// Mitsubishi GX Works2 project: ZhaoQing_HuaCheng1_Debug   PLC: Q06UDEH (continued)

H1000Conveyor7(ConveyorMotor:=H1000Conveyor7IO);
H1000Conveyor7IO.xForward:=M66;
H1000Conveyor7IO.xCWPresent:=X4F;
Y14F:=H1000Conveyor7IO.xMotorCW;
H1000Conveyor7IO.iDeviceID:=1007;

H1000Conveyor8(ConveyorMotor:=H1000Conveyor8IO);
H1000Conveyor8IO.xForward:=M67;
H1000Conveyor8IO.xCWPresent:=X50;
Y150:=H1000Conveyor8IO.xMotorCW;
H1000Conveyor8IO.iDeviceID:=1008;

H1000Conveyor9(ConveyorMotor:=H1000Conveyor9IO);
H1000Conveyor9IO.xForward:=M68;
H1000Conveyor9IO.xCWPresent:=X51;
Y151:=H1000Conveyor9IO.xMotorCW;
H1000Conveyor9IO.iDeviceID:=1009;

H1000Conveyor10(ConveyorMotor:=H1000Conveyor10IO);
H1000Conveyor10IO.xForward:=M67;
H1000Conveyor10IO.xCWPresent:=X52;
Y152:=H1000Conveyor10IO.xMotorCW;
H1000Conveyor10IO.iDeviceID:=1010;
(*注液隔离仓*)
(*FillQuarantineDoorInside(ShuttleCarInOut:= FillQuarantineDoorInsideIO );
FillQuarantineDoorInsideIO.xCylinder:=1;
ShuttleCarCurrentPosition(X109 OR X10A ,X10A ,X109, FALSE,FillQuarantineDoorInsideIO.iCurrentPos);
FillQuarantineDoorInsideIO.xForward:=M191;
FillQuarantineDoorInsideIO.xBackward:=M192 ;
Y160:=FillQuarantineDoorInsideIO.xCW;
Y161:=FillQuarantineDoorInsideIO.xCCW;

FillQuarantineDoorOutside(ShuttleCarInOut:= FillQuarantineDoorOutsideIO );
FillQuarantineDoorOutsideIO.xCylinder:=1;
ShuttleCarCurrentPosition(X10B OR X10C ,X10C ,X10B, FALSE,FillQuarantineDoorOutsideIO.iCurrentPos);
FillQuarantineDoorOutsideIO.xForward:=M193;
FillQuarantineDoorOutsideIO.xBackward:=M194 ;
Y162:=FillQuarantineDoorOutsideIO.xCW;
Y163:=FillQuarantineDoorOutsideIO.xCCW;*)
(*注液入与出线体*)
H850Conveyor1(ConveyorMotor:=H850Conveyor1IO);
H850Conveyor1IO.xForward:=M129;
H850Conveyor1IO.xCWPresent:=X78;
Y178:=H850Conveyor1IO.xMotorCW;
H850Conveyor1IO.iDeviceID:=8501;

H850Conveyor3(ConveyorMotor:=H850Conveyor3IO);
H850Conveyor3IO.xForward:=M130;
H850Conveyor3IO.xCWPresent:=X7A;
Y17A:=H850Conveyor3IO.xMotorCW;
H850Conveyor3IO.iDeviceID:=8503;

H850Conveyor4(ConveyorMotor:=H850Conveyor4IO);
H850Conveyor4IO.xForward:=M131;
H850Conveyor4IO.xCWPresent:=X7B;
Y17B:=H850Conveyor4IO.xMotorCW;
H850Conveyor4IO.iDeviceID:=8504;

H850Conveyor5(ConveyorMotor:=H850Conveyor5IO);
H850Conveyor5IO.xForward:=M132;
H850Conveyor5IO.xCWPresent:=X7C;
Y17C:=H850Conveyor5IO.xMotorCW;
H850Conveyor5IO.iDeviceID:=8505;

H850Conveyor6(ConveyorMotor:=H850Conveyor6IO);
H850Conveyor6IO.xForward:=M133;
H850Conveyor6IO.xCWPresent:=X7D;
Y17D:=H850Conveyor6IO.xMotorCW;
H850Conveyor6IO.iDeviceID:=8506;

H850Conveyor7(ConveyorMotor:=H850Conveyor7IO);
H850Conveyor7IO.xForward:=M164;
H850Conveyor7IO.xCWPresent:=X7E;
Y17E:=H850Conveyor7IO.xMotorCW;
H850Conveyor7IO.iDeviceID:=8507;

H850Rotor(ShuttleCarInOut:=H850RotorIO);
ShuttleCarCurrentPosition(X82 OR X76  ,X82 ,X76, FALSE,H850RotorIO.iCurrentPos);
H850RotorIO.xReady:=TRUE;
H850RotorIO.xForward:=M75;
H850RotorIO.xBackward:=M76;
H850RotorIO.xPosLimit:=X84;
H850RotorIO.xNegLimit:=X85;
Y182:=H850RotorIO.xCW;
Y183:=H850RotorIO.xCCW;
Y1B9:=H850RotorIO.xBrake;

H850RotorConveyor(ConveyorMotor:=H850RotorConveyorIO);
H850RotorConveyorIO.xForward:=M77;
H850RotorConveyorIO.xBackward:=M82;
H850RotorConveyorIO.xCWPresent:=X87;
H850RotorConveyorIO.xCCWPresent:=X86;
Y185:=H850RotorConveyorIO.xMotorCW;
Y184:=H850RotorConveyorIO.xMotorCCW;
H850RotorConveyorIO.xUnloadCCW:=1;
H850RotorConveyorIO.tLoadDelay:=T#2s;
H850RotorConveyorIO.iDeviceID:=8599;

H850Switch(ConveyorEntryIO:=H850SwitchConveyorIn,ConveyorExitIO:=H850SwitchConveyorOut,SwitchIO:=H850SwitchIO);
H850SwitchIO.xLiftCylinderExtendButton:=M71;
H850SwitchIO.xLiftCylinderRetractButton:=M72;
Y189:=H850SwitchIO.xLiftCylinderExtend;
Y188:=H850SwitchIO.xLiftCylinderRetract;
H850SwitchIO.xLiftCylinderExtendDetect:=X88;
H850SwitchIO.xLiftCylinderRetractDetect:=X89;
H850SwitchConveyorIn.xForward:=M70;
H850SwitchConveyorIn.xCWPresent:=XB4;
Y19B:=H850SwitchConveyorIn.xMotorCW;
Y139:=H850SwitchConveyorIn.xMotorCW;(*新加的滚轮电机*)
H850SwitchConveyorIn.tLoadDelay:=T#2s;
H850SwitchConveyorIn.iDeviceID:=8598;
H850SwitchConveyorOut.xForward:=M73;
H850SwitchConveyorOut.xCWPresent:=X8A;
Y18A:=H850SwitchConveyorOut.xMotorCW;
H850SwitchConveyorOut.iDeviceID:=8598;


H850Conveyor8(ConveyorMotor:=H850Conveyor8IO);
H850Conveyor8IO.xForward:=M74;
H850Conveyor8IO.xCWPresent:=X7F;
Y17F:=H850Conveyor8IO.xMotorCW;
H850Conveyor8IO.iDeviceID:=8508;
(*高温库前线体*)
(*-------高温入库分流扫码*)
IF X0BB AND NOT X0BA  THEN 
	Y1BE:=0;
	Y1BF:=1;
END_IF ;
IF ldp(TRUE,X0BA AND D2300=0)  THEN 
	Y1BE:=0;
	Y1BF:=0;
	xscaning1:=1;
END_IF ;
IF ldp(TRUE, D2300=2 OR D2300=3) THEN
	Y1BE:=1;
    Y1BF:=1;
    xscaning1:=0;
END_IF;  
(*阻挡气缸升起，检测有无信号存在，上位机扫码信号复位，可以扫码*)
IF X0BA AND D2300=0 AND Y1BE = 0 AND Y1BF=0 THEN 
	D3300:=2;
END_IF;
(*单体复位后把扫码信息复位*)
IF g_xResetSingle AND g_iDeviceIDSelect=H2200Switch2ConveyorIn.iDeviceID THEN
	xscaning1:=0;
	D3300:=1;
END_IF;
IF D2300 =1 AND g_xReset THEN(*扫码失败复位*)
	D3300:=0;
END_IF;
(* 顶升移载收到物料后复位读码信号*)
(*IF LDP(TRUE,Import1SwitchConveyorOut.xEmpty=0 AND D2300=2) OR LDP(TRUE,Import2SwitchConveyorOut.xEmpty=0 AND D2300=3) THEN*)
	(*修改下复位扫码的时序，分流后再复位扫码信息，方便分流*)
IF( Import1Conveyor1IO.xEmpty=0 AND D2300=2) OR  (Import2Conveyor1IO.xEmpty=0 AND D2300=3) THEN(*效率低*)(*效率低也没办法，分流信息不能提前复位*)
(*IF (Import1SwitchConveyorOut.xBusy AND D2300=2) OR (Import2SwitchConveyorOut.xBusy AND D2300=3) THEN*)
	D3300:=1;    (*接堆垛机那个口顶起来才允许下一次扫码*)(*到达分流顶升移载后复位*)
END_IF;
	(*------高温出库分流扫码*)
	IF X106 THEN 
	xScaning2:=0;
END_IF;
IF X0B9 AND NOT X0B8  THEN 
	Y1BC:=0;
	Y1BD:=1;
END_IF ;
IF X0B8 AND  D2305=0  THEN 
	Y1BC:=0;
	Y1BD:=0;
	xScaning2:=1;
END_IF ;
IF ldp(TRUE,  D2305=2 OR D2305=3) THEN
	Y1BC:=1;
    Y1BD:=1;
    xScaning2:=0;
END_IF;
IF X0B8  AND D2305=0 THEN 
	D3305:=2;
END_IF;
IF X2F OR X39 OR g_xReset THEN(*增加复位信号，扫码失败后按复位按钮*)
	D3305:=1;(*运出之后才允许下一次扫码*)
	END_IF;
(*1巷道入库*)
Import1Conveyor1(ConveyorMotor:=Import1Conveyor1IO);
Import1Conveyor1IO.xForward:=M98;
Import1Conveyor1IO.xCWPresent:=XE3;
Y1F4:=Import1Conveyor1IO.xMotorCW;
Import1Conveyor1IO.iDeviceID:=2290;

Import1Conveyor2(ConveyorMotor:=Import1Conveyor2IO);
Import1Conveyor2IO.tLoadDelay:=T#1s;
Import1Conveyor2IO.xForward:=M99;
Import1Conveyor2IO.xCWPresent:=XE4;
Y1F5:=Import1Conveyor2IO.xMotorCW;
Import1Conveyor2IO.iDeviceID:=2289;

Import1Switch(ConveyorEntryIO:=Import1SwitchConveyorIn,
                          ConveyorExitIO:=Import1SwitchConveyorOut ,
                           SwitchIO:=Import1SwitchIO);
Import1SwitchIO.xLiftCylinderExtendButton:=M147;
Import1SwitchIO.xLiftCylinderRetractButton:=M148;
Import1SwitchIO.xExitBarCylinderRetractButton:=M161;
Y1E0:=Import1SwitchIO.xExitBarCylinderRetract;
Y1E2:=Import1SwitchIO.xLiftCylinderExtend;
Y1E1:=Import1SwitchIO.xLiftCylinderRetract;
Import1SwitchIO.xLiftCylinderExtendDetect:=XE1;
Import1SwitchIO.xLiftCylinderRetractDetect:=XE2; 
Import1SwitchConveyorIn.xCWPresent:=XE0;
Import1SwitchConveyorIn.tLoadDelay:=T#3s;
Import1SwitchConveyorIn.iDeviceID:=2297;
Import1SwitchConveyorOut.xForward:=M149;
Import1SwitchConveyorOut.xCWPresent:=X108;
Y1F6:=Import1SwitchConveyorOut.xMotorCW;
Import1SwitchConveyorOut.iDeviceID:=2297;

Import1LoadCylinder(ShuttleCarInOut:=Import1LoadCylinderIO);
ShuttleCarCurrentPosition(XE7 OR XE6,XE7 ,XE6, FALSE,Import1LoadCylinderIO.iCurrentPos );
Import1LoadCylinderIO.xReady:=TRUE;
Import1LoadCylinderIO.xForward:=M159;
Import1LoadCylinderIO.xBackward:=M160;
Import1LoadCylinderIO.xPosLimit:=TRUE;
Import1LoadCylinderIO.xNegLimit:=TRUE;
Y1E4:=Import1LoadCylinderIO.xCW;
Y1E3:=Import1LoadCylinderIO.xCCW;

(*1巷道出库*)
Export1Conveyor1(ConveyorMotor:=Export1Conveyor1IO);
Export1Conveyor1IO.xForward:=M94;
Export1Conveyor1IO.xCWPresent:=XEC;
Y1F7:=Export1Conveyor1IO.xMotorCW;
Export1Conveyor1IO.iDeviceID:=3081;

Export1Conveyor2(ConveyorMotor:=Export1Conveyor2iO);
Export1Conveyor2IO.xForward:=M95;
Export1Conveyor2IO.xCWPresent:=XEB;
Y1F8:=Export1Conveyor2IO.xMotorCW;
Export1Conveyor2IO.iDeviceID:=3082;

Export1Switch(ConveyorEntryIO:=Export1SwitchConveyorIn,
                          ConveyorExitIO:=Export1SwitchConveyorOut ,
                           SwitchIO:=Export1SwitchIO);
Export1SwitchIO.xLiftCylinderExtendButton:=M150;
Export1SwitchIO.xLiftCylinderRetractButton:=M151;
Y1E7:=Export1SwitchIO.xLiftCylinderExtend;
Y1E6:=Export1SwitchIO.xLiftCylinderRetract;
Export1SwitchIO.xLiftCylinderExtendDetect:=XE9;
Export1SwitchIO.xLiftCylinderRetractDetect:=XEA;
Export1SwitchConveyorIn.xForward:=M152;
Export1SwitchConveyorIn.xCWPresent:=X106;
Export1SwitchConveyorIn.tLoadDelay:=T#2s;
Export1SwitchConveyorIn.iDeviceID:=3083;
Y1F9:=Export1SwitchConveyorIn.xMotorCW;
Export1SwitchConveyorOut.xCWPresent:=X106;
Export1SwitchConveyorOut.iDeviceID:=3083;

Export1LoadCylinder(ShuttleCarInOut:=Export1LoadCylinderIO);
ShuttleCarCurrentPosition(XEF OR XEE ,XEF ,XEE, FALSE,Export1LoadCylinderIO.iCurrentPos);
Export1LoadCylinderIO.xReady:=TRUE;
Export1LoadCylinderIO.xForward:=M157;
Export1LoadCylinderIO.xBackward:=M158;
Export1LoadCylinderIO.xPosLimit:=TRUE;
Export1LoadCylinderIO.xNegLimit:=TRUE;
Y1E9:=Export1LoadCylinderIO.xCW;
Y1E8:=Export1LoadCylinderIO.xCCW;


(*2巷道入库*)
Import2Conveyor1(ConveyorMotor:=Import2Conveyor1IO);
Import2Conveyor1IO.xForward:=M153;
Import2Conveyor1IO.xCWPresent:=XF3;
Y1FA:=Import2Conveyor1IO.xMotorCW;
Import2Conveyor1IO.iDeviceID:=2288;

Import2Conveyor2(ConveyorMotor:=Import2Conveyor2IO);
Import2Conveyor2IO.tLoadDelay:=T#1s;
Import2Conveyor2IO.xForward:=M154;
Import2Conveyor2IO.xCWPresent:=XF4;
Y1FB:=Import2Conveyor2IO.xMotorCW;
Import2Conveyor2IO.iDeviceID:=2287;

Import2Switch(ConveyorEntryIO:=Import2SwitchConveyorIn,
                          ConveyorExitIO:=Import2SwitchConveyorOut ,
                           SwitchIO:=Import2SwitchIO);
Import2SwitchIO.xLiftCylinderExtendButton:=M155;
Import2SwitchIO.xLiftCylinderRetractButton:=M156;
Y1EC:=Import2SwitchIO.xLiftCylinderExtend;
Y1EB:=Import2SwitchIO.xLiftCylinderRetract;
Import2SwitchIO.xLiftCylinderExtendDetect:=XF1;
Import2SwitchIO.xLiftCylinderRetractDetect:=XF2;
Import2SwitchConveyorIn.xCWPresent:=X104;
Import2SwitchConveyorIn.tLoadDelay:=T#2s;
Import2SwitchConveyorIn.iDeviceID:=2296;
Import2SwitchConveyorOut.xForward:=M165;
Import2SwitchConveyorOut.xCWPresent:=X100;
Y1FC:=Import2SwitchConveyorOut.xMotorCW;
Import2SwitchConveyorOut.iDeviceID:=2296;

Import2LoadCylinder(ShuttleCarInOut:=Import2LoadCylinderIO);
ShuttleCarCurrentPosition(XF6 OR XF7 ,XF7 ,XF6, FALSE,Import2LoadCylinderIO.iCurrentPos );
Import2LoadCylinderIO.xReady:=TRUE;
Import2LoadCylinderIO.xForward:=M171;
Import2LoadCylinderIO.xBackward:=M162;
Import2LoadCylinderIO.xPosLimit:=TRUE;
Import2LoadCylinderIO.xNegLimit:=TRUE;
Y1EE:=Import2LoadCylinderIO.xCW;
Y1ED:=Import2LoadCylinderIO.xCCW;

(*2巷道出库*)
Export2Conveyor1(ConveyorMotor:=Export2Conveyor1IO);
Export2Conveyor1IO.xForward:=M96;
Export2Conveyor1IO.xCWPresent:=XFB;
Y1FD:=Export2Conveyor1IO.xMotorCW;
Export2Conveyor1IO.iDeviceID:=3085;

Export2Conveyor2(ConveyorMotor:=Export2Conveyor2iO);
Export2Conveyor2IO.xForward:=M97;
Export2Conveyor2IO.xCWPresent:=XFC;
Y1FE:=Export2Conveyor2IO.xMotorCW;
Export2Conveyor2IO.iDeviceID:=3086;

Export2Switch(ConveyorEntryIO:=Export2SwitchConveyorIn,
                          ConveyorExitIO:=Export2SwitchConveyorOut ,
                           SwitchIO:=Export2SwitchIO);
Export2SwitchIO.xLiftCylinderExtendButton:=M120;
Export2SwitchIO.xLiftCylinderRetractButton:=M121;
Export2SwitchIO.xLiftCylinderExtendInit:=1;
Y1F1:=Export2SwitchIO.xLiftCylinderExtend;
Y1F0:=Export2SwitchIO.xLiftCylinderRetract;
Export2SwitchIO.xLiftCylinderExtendDetect:=XF9;
Export2SwitchIO.xLiftCylinderRetractDetect:=XFA;
Export2SwitchConveyorIn.xForward:=M123;
Export2SwitchConveyorIn.xCWPresent:=X105;
Export2SwitchConveyorIn.tLoadDelay:=T#2s;
Y1FF:=Export2SwitchConveyorIn.xMotorCW;
Export2SwitchConveyorIn.iDeviceID:=3084;
Export2SwitchConveyorOut.xCWPresent:=X105;
Export2SwitchConveyorOut.iDeviceID:=3084;

Export2LoadCylinder(ShuttleCarInOut:=Export2LoadCylinderIO);
ShuttleCarCurrentPosition( XFF OR XFE ,XFF ,XFE, FALSE, Export2LoadCylinderIO.iCurrentPos);
Export2LoadCylinderIO.xReady:=TRUE;
Export2LoadCylinderIO.xForward:=M124;
Export2LoadCylinderIO.xBackward:=M125;
Export2LoadCylinderIO.xPosLimit:=TRUE;
Export2LoadCylinderIO.xNegLimit:=TRUE;
Y1F2:=Export2LoadCylinderIO.xCW;
Y1F3:=Export2LoadCylinderIO.xCCW;




IF g_xAuto THEN
	(**高温库前自动程序**)
	Y1EA:=1;
	m_tonScan2(IN:=xScaning2 ,PT:=T#500ms ,Q:=m_xScan2,ET:= m_tScan2 );(*---------扫码标志位做延时，防止走不到位*)
	Y187:=NOT m_xScan2 AND  m_iExportConveyorOcuppy<>0;(***出库倍速链***)(*---------扫码时停下，扫完走*)
	Y1BA:=NOT m_xScan2 AND  m_iExportConveyorOcuppy<>0;(*后增加滚筒线，在出库线占用状态字有的情况下开始旋转*)
	Y19E :=NOT m_xScan2 AND  m_iExportConveyorOcuppy<>0;
	Y19F:=NOT m_xScan2 AND  m_iExportConveyorOcuppy<>0; 
	(**高温库1巷道出库**)
	(*************************
	上位机通讯程序3
	出口状态  D3105
	1:禁止出库
    2:允许出库
    
    1线堆积(化成线)状态	3106	"1：正常2:堆积 "

2线(二封线)堆积状态	3107	"1：正常2:堆积 "


    收到空框请求D2105
    1：复位，
    2：收到出库请求
	**********************出库********************************)
	(******1巷道******)
	IF NOT XED  AND NOT XEB AND NOT Y1F8 AND Export1LoadCylinderIO.iCurrentPos=2 THEN(*-----这里加了很多条件，保证不会轻易顶起来*)
		D3105:=2;
	ELSE
		D3105:=1;
	END_IF;
	m_tonHangUpChemDalay(IN:= H2200Conveyor5IO.xEmpty=0 OR H2200Conveyor6IO.xEmpty=0  ,PT:=T#30S ,Q:= m_xHangUpChem,ET:= m_tHangUpChemDalayCurrentTime );
	m_tonHangUpPackageDalay(IN:= H3000Conveyor9IO.xEmpty=0 OR H3000Conveyor10IO.xEmpty=0 ,PT:=T#10S ,Q:= m_xHangUpPackage,ET:= m_tHangUpPackageDalayCurrentTime );
	IF m_xHangUpChem THEN
		D3106:=2;
		D3126:=2;
	ELSE
		D3106:=1;
		D3126:=1;
	END_IF;
	
	IF m_xHangUpPackage THEN
		D3107:=2;
		D3127:=2;
	ELSE
		D3107:=1;
		D3127:=1;
	END_IF;
	
	IF D2105=2 THEN
		M883:=1;
	ELSE
		M883:=0;
	END_IF;
	(******2巷道******)
   (*************************
	上位机通讯程序
	出口状态  D3125
	1:禁止出库
    2:允许出库
    1线堆积(化成线)状态	3126	"1：正常2:堆积 "
2线(二封线)堆积状态	3127	"1：正常2:堆积 "

    收到空框请求D2125
    1：复位，
    2：收到出库请求
	**********************出库********************************)
	IF NOT XFD AND Export2LoadCylinderIO.iCurrentPos=2 THEN
		D3125:=2;
	ELSE
		D3125:=1;
	END_IF;
	IF D2125=2 THEN
		M884:=1;
	ELSE
		M884:=0;
	END_IF;
	(*********************入库****************************)
	(***********************************
	入口状态 D3100
	1:无电池入库请求
     2:有电池入库请求
	************************************)
	(******1巷道******)
	m_tonImport1RequestDalay(IN:= XE5 ,PT:= t#3S ,Q:= m_xImport1RequestDalay ,ET:=m_tImport1RequestDalaDalayCurren);
	IF m_xImport1RequestDalay AND Import1LoadCylinderIO.iCurrentPos=2 THEN
		D3100:=2;
	ELSE
		D3100:=1;
    END_IF;  
    (******2巷道******)
	m_tonImport2RequestDalay(IN:= XF5 ,PT:= t#3S ,Q:= m_xImport2RequestDalay ,ET:=m_tImport2RequestDalaDalayCurren);    
    IF m_xImport2RequestDalay  AND Import2LoadCylinderIO.iCurrentPos=2 THEN
		D3120:=2;
	ELSE
		D3120:=1;
    END_IF;
    (*******************************************************)
    (******高温出库分流******)
    (***********************************
	有板状态 D3305
	1：无板，2：有板
    分流方向 D2305
0：复位
1：读码失败
2：满筐进加压化成
3：满筐进二封
4：空筐回流进注液
	************************************)
	(*IF H3000SwitchPackageConveyorIn.xEmpty=0 THEN
		D3305:=1;
	ELSE
		D3305:=2;
	END_IF;*)
	IF D2305=2 THEN
		M882:=1;
	END_IF;
	IF D2305 =3 THEN
		M882:=0;
	END_IF;
	(**********************************)
	 (******高温出库后升降机2分流******)
	     (***********************************
	有板状态 D3310
	1：无板，2：有板
    分流方向 D2310
0：复位
1：读码失败
2：空筐去注液
3：满筐去加压化成
	************************************)
	IF X3B THEN
		D3310:=2;
	ELSE
		D3310:=1;
	END_IF;
	(*
	IF D2310=2 THEN        ------------这段屏蔽了，直接加到xcondition里了
        Lifter2ExportChem:=01;
	END_IF;
	IF D2310=3 THEN
        Lifter2ExportChem:=1;
	END_IF;
	*)
	(*************	"化成后站台40082335	5	
	分流方向	2335	"0：复位
1：读码失败
2：处理完成放行"
"**********************)



	IF H1000Conveyor2IO.xEmpty=0 THEN
		D3335:=2;
	ELSE
		D3335:=1;
	END_IF;
	IF NOT H850Conveyor8IO.xEmpty THEN
		D3340:=2;
	ELSE
		D3340:=1;
		END_IF;
  (***********************************)
	IF  LDP(TRUE,M883) AND XED THEN
        Export1LoadCylinderIO.xMDIExe:=1;
        Export1LoadCylinderIO.iDestinationPos:=1;
	END_IF;
	IF NOT XED AND NOT XEB  AND NOT Y1F8 AND  Export1Conveyor2IO.xEmpty AND NOT Export1Conveyor2IO.xBusy THEN
        Export1LoadCylinderIO.xMDIExe:=1;
        Export1LoadCylinderIO.iDestinationPos:=2;
     END_IF;		
	Export1Conveyor2IO.xLoad:=XED AND Export1LoadCylinderIO.iCurrentPos=1;
	Export1Conveyor2IO.xUnload:=Export1Conveyor1IO.xEmpty;
	Export1Conveyor1IO.xLoad:=Export1Conveyor2IO.xNextRun;

	Export1Conveyor1Io.xUnload:=Export1SwitchConveyorIn.xEmpty  AND  m_iExportConveyorOcuppy=1 AND  NOT M173;
	IF Export1Conveyor1Io.xEmpty=0 AND m_xExportConveyorIdle THEN
		m_iExportConveyorOcuppy:=1;
	END_IF;
	Export1SwitchIO.xEntryEnable:=Export1Conveyor1Io.xNextRun;
	Export1SwitchIO.xSwithEnable:=1;
	(*倍速链上只有一个物料出库*)
   Export1SwitchIO.xExitEnable:=(H3000SwitchChemConveyorIn.xEmpty AND M882) OR (H3000Conveyor1IO.xEmpty AND NOT M882);
	(**高温库2巷道出库**)
	IF  LDP(TRUE,M884) AND XFD THEN
        Export2LoadCylinderIO.xMDIExe:=1;
        Export2LoadCylinderIO.iDestinationPos:=1;
	END_IF;
	IF NOT XFD  AND NOT Export2Conveyor1IO.xBusy AND Export2Conveyor1IO.xEmpty  THEN
        Export2LoadCylinderIO.xMDIExe:=1;
        Export2LoadCylinderIO.iDestinationPos:=2;
     END_IF;	
	Export2Conveyor1IO.xLoad:=XFD AND Export2LoadCylinderIO.iCurrentPos=1;
	Export2Conveyor1IO.xUnload:=Export2Conveyor2IO.xEmpty;
	Export2Conveyor2IO.xLoad:=Export2Conveyor1IO.xNextRun;
(*	Export2Conveyor2Io.xUnload:=Export2SwitchConveyorIn.xEmpty AND NOT XE8 AND NOT Y1E5;(*增加阻挡器信号与到位信号*)
	Export2Conveyor2Io.xUnload:=Export2SwitchConveyorIn.xEmpty AND  m_iExportConveyorOcuppy=2 AND NOT M173;
	Export2SwitchIO.xEntryEnable:=Export2Conveyor2Io.xNextRun;
	Export2SwitchIO.xSwithEnable:=1;

	IF Export2Conveyor2Io.xEmpty=0 AND m_xExportConveyorIdle  THEN
		m_iExportConveyorOcuppy:=2;
	END_IF;
	IF m_iExportConveyorOcuppy=2  THEN
		Y1E5:=1;(*1巷道出库阻挡器*)
		Export1SwitchIO.xLiftCylinderExtendInit:=0;
	ELSE
		Y1E5:=0;(*1巷道出库阻挡器*)
		Export1SwitchIO.xLiftCylinderExtendInit:=1;	
	END_IF;
	
	Export2SwitchIO.xExitEnable:=(H3000SwitchChemConveyorIn.xEmpty AND M882) OR (H3000Conveyor1IO.xEmpty AND NOT M882);
	(*占用信号的复位*)
	IF LDP(TRUE,H3000SwitchChemConveyorIn.xEmpty=0 AND M882) OR LDP(TRUE,H3000Conveyor1IO.xEmpty=0 AND NOT M882) THEN
		m_iExportConveyorOcuppy:=0;
	END_IF;
	
	m_tonExportConveyorOcuppy(IN:= m_iExportConveyorOcuppy=0 ,PT:= T#3s ,Q:= m_xExportConveyorIdle ,ET:= m_tExportConveyorOcuppyCurrent );

	(*满框出库去二次封装线体*)
	H3000SwitchQuadPackageIO.xEntryEnable:=1;(*这里要加扫码条件*)
	H3000SwitchQuadPackageIO.xSwithEnable:= NOT M882;(*触摸屏上按钮选择去化成还是去二封，后期通过上位机扫码给出*)
	IF H3000SwitchQuadPackageIO.xSwithEnable THEN
		H3000SwitchQuadPackageio.xExitEnable:=H3000Conveyor1IO.xEmpty;
		H3000Conveyor1Io.xLoad:=H3000SwitchPackageConveyorOut.xNextRun;
	ELSE
		H3000SwitchQuadPackageio.xExitEnable:=0;	
		H3000Conveyor1Io.xLoad:=0;
	END_IF;
	H3000Conveyor1IO.xUnload:=H3000Conveyor2IO.xEmpty;
	H3000Conveyor2IO.xLoad:=H3000Conveyor1IO.xNextRun;
	H3000Conveyor2IO.xUnload:=H3000Conveyor3IO.xEmpty;
	H3000Conveyor3IO.xLoad:=H3000Conveyor2IO.xNextRun;	
	H3000Conveyor3IO.xUnload:=H3000Conveyor4IO.xEmpty;
	H3000Conveyor4IO.xLoad:=H3000Conveyor3IO.xNextRun;
	H3000Conveyor4IO.xUnload:=H3000Conveyor5IO.xEmpty;
	H3000Conveyor5IO.xLoad:=H3000Conveyor4IO.xNextRun;
	H3000Conveyor5IO.xUnload:=H3000Conveyor6IO.xEmpty;
	H3000Conveyor6IO.xLoad:=H3000Conveyor5IO.xNextRun;
	H3000Conveyor6IO.xUnload:=H3000Conveyor7IO.xEmpty;
	H3000Conveyor7IO.xLoad:=H3000Conveyor6IO.xNextRun;
	H3000Conveyor7IO.xUnload:=H3000Conveyor8IO.xEmpty;
	H3000Conveyor8IO.xLoad:=H3000Conveyor7IO.xNextRun;	
	H3000Conveyor8IO.xUnload:=H3000Conveyor9IO.xEmpty;
	H3000Conveyor9IO.xLoad:=H3000Conveyor8IO.xNextRun;	
	H3000Conveyor9IO.xUnload:=H3000Conveyor10IO.xEmpty;
	H3000Conveyor10IO.xLoad:=H3000Conveyor9IO.xNextRun;
	H3000Conveyor10IO.xUnload:=D401.0;
	D201.0:=H3000Conveyor10IO.xNextRun;
    (**满框去化成**)
	H3000SwitchChemIO.xEntryEnable:=1;
	H3000SwitchChemIO.xSwithEnable:=1;
	H3000SwitchChemIO.xExitEnable:=H3000ChemConveyor2IO.xEmpty;
	H3000SwitchPackageConveyorIn.xUnload:=H3000SwitchChemConveyorIn.xEmpty;
	H3000ChemConveyor2IO.xLoad:=H3000SwitchChemConveyorOut.xNextRun;
	H3000ChemConveyor2IO.xUnload:=H3000ChemConveyor3IO.xEmpty;
	H3000ChemConveyor3IO.xLoad:=H3000ChemConveyor2IO.xNextRun;
	(*临时程序，Lifter2ExportChem:=1;以后要考虑空框回注液的程序，上位机扫码后判断是满框去化成还是空框去注液*)
	IF H3000ChemConveyor3IO.xEmpty=0 AND ( Lifter2TaskID=3 OR Lifter2TaskID=4)  THEN(*这里加扫码成功条件*)
		Lifter2IO.xMDIExe:=1;
		Lifter2IO.iDestinationPos:=5;
	END_IF;
	IF Lifter2IO.iCurrentPos=5 AND abs(D190-Lifter2Position[Lifter2IO.iDestinationPos])<20 AND (Lifter2TaskID=3 OR Lifter2TaskID=4)   THEN	
        Conveyor2IO.xLoad:=H3000ChemConveyor3IO.xNextRun;
        H3000ChemConveyor3IO.xUnload:=Conveyor2IO.xEmpty AND H2200Conveyor1io.xEmpty;(*-------这里防止东西堵在车上*)
         Conveyor2IO.xloadCCW:=0;
	ELSE
		H3000ChemConveyor3IO.xUnload:=0;
	END_IF; 
	   IF Conveyor2IO.xEmpty=0 AND Lifter2TaskID=3 THEN
	   		Lifter2IO.xMDIExe:=1;
			Lifter2IO.iDestinationPos:=4;
	   END_IF;
	   	   IF Conveyor2IO.xEmpty=0 AND Lifter2TaskID=4 THEN
	   		Lifter2IO.xMDIExe:=1;
			Lifter2IO.iDestinationPos:=3;
	   END_IF;
	 IF Lifter2IO.iCurrentPos=4 AND abs(D190-Lifter2Position[Lifter2IO.iDestinationPos])<=20  THEN	
	 	H2200Conveyor1IO.xLoad:=Conveyor2IO.xNextRun; 
	 	Conveyor2IO.xUnload:=H2200Conveyor1IO.xEmpty;
	 	Conveyor2IO.xUnloadCCW:=0;
	 ELSE
	 	H2200Conveyor1IO.xLoad:=0;
	 END_IF;  
	      
	H2200Conveyor1IO.xUnload:=H2200Conveyor2IO.xEmpty;
	H2200Conveyor2IO.xLoad:=H2200Conveyor1IO.xNextRun;
	H2200Conveyor2IO.xUnload:=H2200Conveyor3IO.xEmpty;
	H2200Conveyor3IO.xLoad:=H2200Conveyor2IO.xNextRun;	
	H2200Conveyor3IO.xUnload:=H2200Conveyor4IO.xEmpty;
	H2200Conveyor4IO.xLoad:=H2200Conveyor3IO.xNextRun;
	H2200Conveyor4IO.xUnload:=H2200Conveyor5IO.xEmpty;
	H2200Conveyor5IO.xLoad:=H2200Conveyor4IO.xNextRun;
	H2200Conveyor5IO.xUnload:=H2200Conveyor6IO.xEmpty;
	H2200Conveyor6IO.xLoad:=H2200Conveyor5IO.xNextRun;
	H2200Conveyor6IO.xUnload:=H2200Conveyor7IO.xEmpty;
	H2200Conveyor7IO.xLoad:=H2200Conveyor6IO.xNextRun;
	H2200Conveyor7IO.xUnload:=H2200Conveyor8IO.xEmpty;
	H2200Conveyor8IO.xLoad:=H2200Conveyor7IO.xNextRun;	
	H2200Conveyor8IO.xUnload:=H2200Conveyor9IO.xEmpty;
	H2200Conveyor9IO.xLoad:=H2200Conveyor8IO.xNextRun;	
	H2200Conveyor9IO.xUnload:=H2200Conveyor10IO.xEmpty;
	H2200Conveyor10IO.xLoad:=H2200Conveyor9IO.xNextRun;
	H2200Conveyor10IO.xUnload:=D401.1;
	D201.1:=H2200Conveyor10IO.xNextRun;
	(*化成回流线体*)
	D201.2:=H1000Conveyor10IO.xEmpty;
	H1000Conveyor10IO.xLoad:=D401.2;
	H1000Conveyor10IO.xUnload:=H1000Conveyor9IO.xEmpty;
    H1000Conveyor9IO.xLoad:=H1000Conveyor10IO.xNextRun;
    H1000Conveyor9IO.xUnload:=H1000Conveyor8IO.xEmpty;
    H1000Conveyor8IO.xLoad:=H1000Conveyor9IO.xNextRun;
    H1000Conveyor8IO.xUnload:=H1000Conveyor7IO.xEmpty;
    H1000Conveyor7IO.xLoad:=H1000Conveyor8IO.xNextRun;
    H1000Conveyor7IO.xUnload:=H1000Conveyor6IO.xEmpty;
    H1000Conveyor6IO.xLoad:=H1000Conveyor7IO.xNextRun;
    H1000Conveyor6IO.xUnload:=H1000Conveyor5IO.xEmpty;
    H1000Conveyor5IO.xLoad:=H1000Conveyor6IO.xNextRun;
    H1000Conveyor5IO.xUnload:=H1000Conveyor4IO.xEmpty;
    H1000Conveyor4IO.xLoad:=H1000Conveyor5IO.xNextRun;
    H1000Conveyor4IO.xUnload:=H1000Conveyor3IO.xEmpty;
    H1000Conveyor3IO.xLoad:=H1000Conveyor4IO.xNextRun;
    H1000Conveyor3IO.xUnload:=H1000Conveyor2IO.xEmpty;
    H1000Conveyor2IO.xLoad:=H1000Conveyor3IO.xNextRun;  
    H1000Conveyor2IO.xUnload:=H1000Conveyor1IO.xEmpty AND D2335=2;(*------这里加个条件，H1000右边扫码位置*)
    H1000Conveyor1IO.xLoad:=H1000Conveyor2IO.xNextRun; 
    IF H1000Conveyor1IO.xEmpty=0 AND Lifter2TaskID=2 THEN
    	Lifter2IO.xMDIExe:=1;
    	Lifter2IO.iDestinationPos:=2;
    END_IF;    
    IF Lifter2IO.iCurrentPos=2 AND abs(D190-Lifter2Position[Lifter2IO.iDestinationPos])<20 AND Lifter2TaskID=2  THEN (*-------这里改成了20*)
    	H1000Conveyor1IO.xUnload:=Conveyor2IO.xEmpty;
     	Conveyor2IO.xLoad:=H1000Conveyor1IO.xNextRun;     	
    	Conveyor2IO.xloadCCW:=1;
    ELSE
    	H1000Conveyor1IO.xUnload:=0;
    END_IF;
   (*========================================================*)
   (*注液RGV*)
    (*  FillingStab1.xLoadRequest:=X80;*)(*空框上料*)
   (*   FillingStab1.xUnloadRequest:=X81;*)(*满框下料*)
   (*    Y180:= FillingStab1.xLoadRequestAkn;(*空框上料完成*)
    (*   Y181:= FillingStab1.xUnloadRequestAkn;(*满框下料完成*)
       
     (*  FillingStab2.xLoadRequest:=X82;(*空框上料*)
     (*  FillingStab2.xUnloadRequest:=X83;(*满框下料*) 
    (*    Y182:=FillingStab2.xLoadRequestAkn;(*空框上料完成*)
    (*    Y183:=FillingStab2.xUnloadRequestAkn; (*满框下料完成*)   
    
   (*     FillingStab3.xLoadRequest:=X82;(*空框上料*)
     (*  FillingStab3.xUnloadRequest:=X83;(*满框下料*) 
    (*    Y182:=FillingStab3.xLoadRequestAkn;(*空框上料完成*)
  (*      Y183:=FillingStab3.xUnloadRequestAkn; (*满框下料完成*)        
  
      (*     FillingStab4.xLoadRequest:=X82;(*空框上料*)
     (*  FillingStab4.xUnloadRequest:=X83;(*满框下料*) 
    (*    Y182:=FillingStab4.xLoadRequestAkn;(*空框上料完成*)
  (*      Y183:=FillingStab4.xUnloadRequestAkn; (*满框下料完成*)           
	(*发送*)
   D241:=FillingRGV.iDestinationPos;	
   D242.0:=FillingRGV.xAuto; 	
   D242.1:=FillingRGV.xMdiExe;
   D242.2:=FillingRGV.xLoad1;
   D242.3:=FillingRGV.xUnload1;
   D242.4:=FillingStab1.xLoadRequest;
   D242.5:=FillingStab2.xLoadRequest;
   D242.6:=FillingStab3.xLoadRequest;
   D242.7:=FillingStab4.xLoadRequest;
   D242.8:=FillingStab1.xUnloadRequest;
   D242.9:=FillingStab2.xUnloadRequest;
   D242.A:=FillingStab3.xUnloadRequest;
   D242.B:=FillingStab4.xUnloadRequest;
   D244.C:=H850Conveyor1IO.xEmpty;
   D244.D:=H850Conveyor1IO.xNextRun;
   D244.E:=H850Conveyor4IO.xEmpty; 
     
   D243.0:=FillingRGV.xRemoteReset;

   FillingRGV.xRemoteReset:=M178;
   FillingRGV.xAuto:=M179;
   (*接收*)
    FillingRGV.iCurrentPostion:=D441;
   FillingStab1.xLoadRequestAkn:=D442.0;
   FillingStab2.xLoadRequestAkn:=D442.1;
   FillingStab3.xLoadRequestAkn:=D442.2;
  FillingStab4.xLoadRequestAkn:=D442.3;
  FillingStab1.xUnloadRequestAkn:=D442.4;
   FillingStab2.xUnloadRequestAkn:= D442.5;
   FillingStab3.xUnloadRequestAkn:= D442.6; 
   FillingStab4.xUnloadRequestAkn:= D442.7; 
	H850Conveyor1IO.xUnload:=D442.8;
	H850Conveyor4IO.xLoad:=D442.9;
   FillingRGV.xCollisionAlarm:=D443.0;

      (*去空框上下料位置*)(*满框上下料位置*)
    IF M180 THEN
   	FillingRGV.xMdiExe:=1;
   	FillingRGV.iDestinationPos:=7;
    END_IF;   
      (*1号注液机满框下料*) 
   IF M181 THEN
   	FillingRGV.xMdiExe:=1;
   	FillingRGV.iDestinationPos:=1;
   END_IF;
    IF M182 THEN
   	FillingRGV.xMdiExe:=1;
   	FillingRGV.iDestinationPos:=2;
   END_IF;        
      (*2号注液机*) 
   IF M183 THEN
   	FillingRGV.xMdiExe:=1;
   	FillingRGV.iDestinationPos:=3;
   END_IF;  
   IF M184 THEN
   	FillingRGV.xMdiExe:=1;
   	FillingRGV.iDestinationPos:=4;
   END_IF;         
       (*3号注液机*) 
   IF M185 THEN
   	FillingRGV.xMdiExe:=1;
   	FillingRGV.iDestinationPos:=5;
   END_IF;  
   IF M186 THEN
   	FillingRGV.xMdiExe:=1;
   	FillingRGV.iDestinationPos:=6;
   END_IF;  
       (*4号注液机*) 
   IF M187 THEN
   	FillingRGV.xMdiExe:=1;
   	FillingRGV.iDestinationPos:=8;
   END_IF;  
   IF M188 THEN
   	FillingRGV.xMdiExe:=1;
   	FillingRGV.iDestinationPos:=9;
   END_IF;  
   
    (*========================================================*)
	(*注液设备满框入库*)
	H850Conveyor4IO.xLoad:=(M880 OR XD9) AND NOT M172;(*-----加了个按钮*)(*m172,禁止注液上料*)
	H850Conveyor4IO.xUnload:=H850Conveyor5IO.xEmpty;
	H850Conveyor5IO.xLoad:=H850Conveyor4IO.xNextRun;
	H850Conveyor5IO.xUnload:=H850Conveyor6IO.xEmpty;
        IF ldp(TRUE,  H850Conveyor6IO.xEmpty=0) THEN
    		D10:=D10+1;
    	END_IF;
    	(*清零程序*)
    	IF M126 THEN
    		D10:=0;
    	END_IF;
	H850Conveyor6IO.xLoad:=H850Conveyor5IO.xNextRun;	
	IF H850RotorConveyorIO.xEmpty THEN
		 H850RotorIO.xMDIExe:=1;
		  H850RotorIO.iDestinationPos:=1;
	END_IF;
	IF H850RotorConveyorIO.xEmpty=0 THEN                    
		 H850RotorIO.xMDIExe:=1;
		  H850RotorIO.iDestinationPos:=2;
	END_IF;	
	IF H850RotorIO.iCurrentPos=1 THEN
    H850Conveyor6IO.xUnload:=H850RotorConveyorIO.xEmpty;
	ELSE
	 H850Conveyor6IO.xUnload:=0;
	END_IF;	
	H850RotorConveyorIO.xLoad:=H850Conveyor6IO.xNextRun;
	IF H850RotorIO.iCurrentPos=2 THEN
		H850RotorConveyorIO.xUnload:=H850SwitchConveyorIn.xEmpty AND H850SwitchConveyorOut.xEmpty;
	ELSE
		H850RotorConveyorIO.xUnload:=0;
	END_IF;
	H850SwitchIO.xEntryEnable:=H850RotorConveyorIO.xNextRun;	
	H850SwitchIO.xSwithEnable:=1;
	H850SwitchIO.xExitEnable:=H850Conveyor7IO.xEmpty;
    H850Conveyor7IO.xLoad:=H850SwitchConveyorOut.xNextRun;
    
    H850Conveyor7IO.xUnload:=H850Conveyor8IO.xEmpty;
    H850Conveyor8IO.xLoad:=H850Conveyor7IO.xNextRun;
    
    IF H850Conveyor8IO.xEmpty=0 AND Lifter2TaskID=1 THEN
    	Lifter2IO.xMDIExe:=1;
    	Lifter2IO.iDestinationPos:=1;
    END_IF;
    IF Lifter2IO.iCurrentPos=1 AND ABS(D190-Lifter2Position[Lifter2IO.iDestinationPos])<20 THEN(*--------改成了20*)
    	H850Conveyor8IO.xUnload:= Conveyor2IO.xEmpty AND Lifter2TaskID=1;(*--------这里加了task条件，不会无条件进升降机了*)
    	Conveyor2IO.xLoad:=H850Conveyor8IO.xNextRun;
        Conveyor2IO.xloadCCW:=0;
    ELSE
    	H850Conveyor8IO.xUnload:=0;
    END_IF;
     IF (Lifter2TaskID=1 OR Lifter2TaskID=2 OR Lifter2TaskID=4) AND Conveyor2IO.xEmpty=0 THEN(*只要不是加压化成的 满框都要入库*)(*这里加扫码条件*)
     	Lifter2IO.xMDIExe:=1;
    	Lifter2IO.iDestinationPos:=3;
     END_IF;
    IF Lifter2IO.iCurrentPos=3 AND ABS(D190-Lifter2Position[Lifter2IO.iDestinationPos])<20 THEN	 (*-------这里改成了20*)
		Conveyor2IO.xUnload:=H2200ImportConveyor2IO.xEmpty;
		H2200ImportConveyor2IO.xLoad:=Conveyor2IO.xNextRun;  
		Conveyor2IO.xUnloadCCW:=1;
    ELSE
    	 H2200ImportConveyor2IO.xLoad:=0; 	
    END_IF;
    (*不在目标位置不可上下料*)
    IF ABS(D190-Lifter2Position[Lifter2IO.iDestinationPos])>20 
    	OR  LIfter2IO.iCurrentPos=5 
    	OR LIfter2IO.iCurrentPos=1 
    	OR Lifter2IO.iCurrentPos=2   THEN (*-------这里改成了20,和1层2层5层不准下*)
    	Conveyor2IO.xUnload:=0;
    END_IF;
    IF ABS(D190-Lifter2Position[Lifter2IO.iDestinationPos])>20 
    	OR Lifter2IO.iCurrentPos=3
    	OR Lifter2IO.iCurrentPos=4 THEN
    	Conveyor2IO.xLoad:=0;
    END_IF;
    
    H2200ImportConveyor2IO.xUnload:=H2200ImportConveyor3IO.xEmpty;
    H2200ImportConveyor3IO.xLoad:=H2200ImportConveyor2IO.xNextRun;
    
    (*满框入库任务*)
    IF H2200Switch1TaskID=5 THEN
	    H2200ImportConveyor3IO.xUnload:= H2200ImportConveyor1IO.xEmpty AND H2200Switch1ConveyorOut.xEmpty;
	    H2200Switch1ConveyorOut.xLoad:=H2200ImportConveyor3IO.xNextRun; 
	    H2200Switch1IO.xLiftCylinderExtendInit:=1;	          	    
    ELSE
    	 H2200ImportConveyor3IO.xUnload:=0;
    	 
    END_IF;
    H2200Switch1ConveyorOut.xUnload:=H2200ImportConveyor1IO.xEmpty AND H2200Switch1TaskID=5 ; 
    H2200ImportConveyor1IO.xLoad:=H2200Switch1ConveyorOut.xNextRun;
    H2200ImportConveyor1IO.xUnload:=H2200Switch2ConveyorIn.xEmpty;
    H2200Switch2IO.xEntryEnable:=H2200ImportConveyor1IO.xNextRun;
    H2200Switch2IO.xSwithEnable:=1;
    (*-----此处有挡停后要加挡停条件，还要把巷道2的为空的条件加上,已经加上读码条件来互锁入库传输线*)
    H2200Switch2IO.xExitEnable:=( Import1SwitchConveyorIn.xEmpty AND D2300=2) (*扫码后*)
                                                        OR ( Import2SwitchConveyorIn.xEmpty AND D2300=3) 
                                                        OR D2300=0(*未扫码*)
                                                        OR D2300=1(*扫码失败*)
                                                        OR X0BA ;(*扫码开关*)
    (*1巷道入库*)
    Import1SwitchIO.xEntryEnable:=D2300>1;
    Import1SwitchIO.xSwithEnable:=D2300=2 ;(*临时程序*)
    Import1SwitchIO.xExitEnable:=(Import1Conveyor1IO.xEmpty AND D2300=2) OR (Import2SwitchConveyorIn.xEmpty AND D2300=3) ;
    Import1Conveyor1IO.xLoad:=Import1SwitchConveyorOut.xNextRun;
    Import1Conveyor1IO.xUnload:=Import1Conveyor2IO.xEmpty AND NOT XE5;
    Import1Conveyor2IO.xLoad:=Import1Conveyor1IO.xNextRun;
    
    IF Import1Conveyor2IO.xEmpty=0 AND XE5 THEN
    	Import1LoadCylinderIO.xMDIExe:=1;
    	Import1LoadCylinderIO.iDestinationPos:=2;
    	Import1Conveyor2IO.xPutInto:=0;
    END_IF;
    IF NOT XE5 THEN
    	Import1LoadCylinderIO.xMDIExe:=1;
    	Import1LoadCylinderIO.iDestinationPos:=1;	
    END_IF;
    IF LDP(TRUE, Import1LoadCylinderIO.iCurrentPos=1) THEN
    	Import1Conveyor2IO.xPutInto:=1;
    END_IF;
 (*2巷道入库*)
     Import2SwitchIO.xEntryEnable:=1;
    Import2SwitchIO.xSwithEnable:=1;
    Import2SwitchIO.xExitEnable:=Import2Conveyor1IO.xEmpty;
    Import2Conveyor1IO.xLoad:=Import2SwitchConveyorOut.xNextRun;
    Import2Conveyor1IO.xUnload:=Import2Conveyor2IO.xEmpty AND NOT XF5;
    Import2Conveyor2IO.xLoad:=Import2Conveyor1IO.xNextRun;